   "EMS".Carrier[78].SDC_OUT.HeartBeat := "Clock_1Hz";
   "EMS".Carrier[79].SDC_OUT.HeartBeat := "Clock_1Hz";
   "EMS".Carrier[80].SDC_OUT.HeartBeat := "Clock_1Hz";
END_REGION

REGION Network 2
   // **********************************************************************************************************************
   // 
   // Carrier 71 I-Device Data Transfer Interlocks from Carrier to SDC
   // 
   // **********************************************************************************************************************
   RUNG wire#powerrail
      Coil( "SectionComment" )
   END_RUNG
   // the same network as SCL:
   "SectionComment" := TRUE;
END_REGION

REGION Network 3
   RUNG wire#powerrail
      Contact( "Carrier_71_Status.0" )
      Coil( "EMS".Carrier[71].SDC_IN.HeartBeat )
   END_RUNG
   // the same network as SCL:
   "EMS".Carrier[71].SDC_IN.HeartBeat := "Carrier_71_Status.0";
END_REGION

REGION Network 4
   "C71_Heartbeat_On_Timer".TON(IN := "EMS".Carrier[71].SDC_IN.HeartBeat, PT := T#3s);
END_REGION

REGION Network 5
   "C71_Heartbeat_Off_Timer".TON(IN := NOT "EMS".Carrier[71].SDC_IN.HeartBeat, PT := T#3s);
END_REGION

REGION Network 6
   RUNG wire#powerrail
      Contact( "Carrier_71_Status.7" )
      wire#w1
      Coil( "EMS".Carrier[71].CommFlt )
   END_RUNG
   RUNG wire#powerrail
      Contact( "C71_Heartbeat_On_Timer".Q )
   END_RUNG wire#w1
   RUNG wire#powerrail
      Contact( "C71_Heartbeat_Off_Timer".Q )
   END_RUNG wire#w1
   // the same network as SCL:
   "EMS".Carrier[71].CommFlt := "Carrier_71_Status.7" OR "C71_Heartbeat_On_Timer".Q OR "C71_Heartbeat_Off_Timer".Q;
END_REGION

REGION Network 7
   RUNG wire#powerrail
      Contact( "EMS".Carrier[71].CommFlt )
      JumpCoil( C71_Comm_Fault )
   END_RUNG
   // the same network as SCL:
   IF "EMS".Carrier[71].CommFlt THEN GOTO C71_Comm_Fault; END_IF;
END_REGION

REGION Network 8
   RUNG wire#powerrail
      { S7_Templates := "SrcType := Word" } NE_Contact(in1 := "Carrier_71_CarrierNumber", in2 := 0)
      Move(in := "Carrier_71_CarrierNumber", out1 => "EMS".Carrier[71].SDC_IN.CarrierNumber)
   END_RUNG
   // the same network as SCL:
   IF "Carrier_71_CarrierNumber" <> 0 THEN
       "EMS".Carrier[71].SDC_IN.CarrierNumber := "Carrier_71_CarrierNumber";
   END_IF;
END_REGION

REGION Network 9
   RUNG wire#powerrail
      { S7_Templates := "SrcType := DWord" } NE_Contact(in1 := "Carrier_71_CarrierPosition", in2 := 0)
      Move(in := "Carrier_71_CarrierPosition", out1 => "EMS".Carrier[71].SDC_IN.CarrierPosition)
   END_RUNG
   // the same network as SCL:
   IF "Carrier_71_CarrierPosition" <> 0 THEN
       "EMS".Carrier[71].SDC_IN.CarrierPosition := "Carrier_71_CarrierPosition";
   END_IF;
END_REGION

REGION Network 10
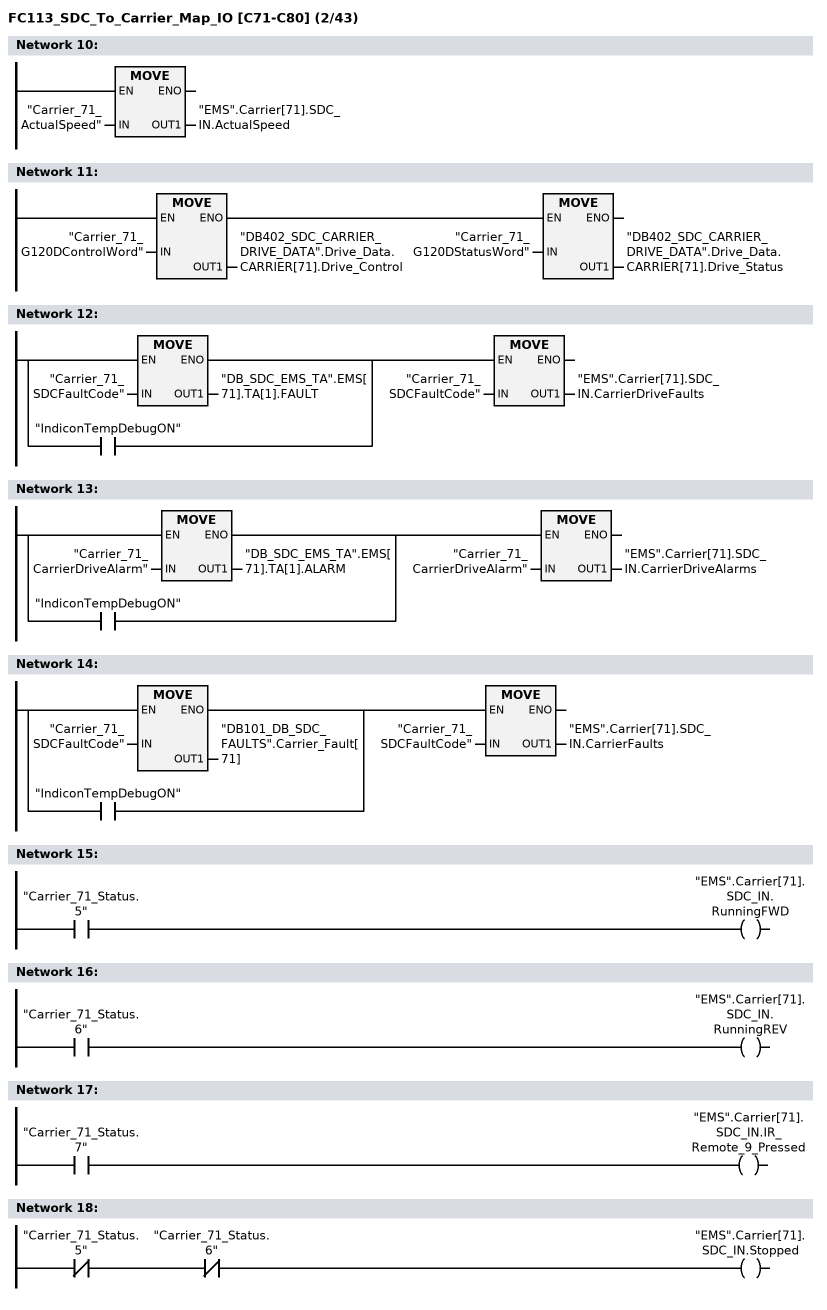
   RUNG wire#powerrail
      Move(in := "Carrier_71_ActualSpeed", out1 => "EMS".Carrier[71].SDC_IN.ActualSpeed)
   END_RUNG
   // the same network as SCL:
   "EMS".Carrier[71].SDC_IN.ActualSpeed := "Carrier_71_ActualSpeed";
END_REGION

REGION Network 11
   RUNG wire#powerrail
      Move(in := "Carrier_71_G120DControlWord", out1 => "DB402_SDC_CARRIER_DRIVE_DATA".Drive_Data.CARRIER[71].Drive_Control)
      Move(in := "Carrier_71_G120DStatusWord", out1 => "DB402_SDC_CARRIER_DRIVE_DATA".Drive_Data.CARRIER[71].Drive_Status)
   END_RUNG
   // the same network as SCL:
   "DB402_SDC_CARRIER_DRIVE_DATA".Drive_Data.CARRIER[71].Drive_Control := "Carrier_71_G120DControlWord";
   "DB402_SDC_CARRIER_DRIVE_DATA".Drive_Data.CARRIER[71].Drive_Status := "Carrier_71_G120DStatusWord";
END_REGION

REGION Network 12
   RUNG wire#powerrail
      Move(in := "Carrier_71_SDCFaultCode", out1 => "DB_SDC_EMS_TA".EMS[71].TA[1].FAULT)
      wire#w1
      Move(in := "Carrier_71_SDCFaultCode", out1 => "EMS".Carrier[71].SDC_IN.CarrierDriveFaults)
   END_RUNG
   RUNG wire#powerrail
      Contact( "IndiconTempDebugON" )
   END_RUNG wire#w1
   // the same network as SCL:
   "DB_SDC_EMS_TA".EMS[71].TA[1].FAULT := "Carrier_71_SDCFaultCode";
   IF TRUE OR "IndiconTempDebugON" THEN
       "EMS".Carrier[71].SDC_IN.CarrierDriveFaults := "Carrier_71_SDCFaultCode";
   END_IF;
END_REGION

REGION Network 13
   RUNG wire#powerrail
      Move(in := "Carrier_71_CarrierDriveAlarm", out1 => "DB_SDC_EMS_TA".EMS[71].TA[1].ALARM)
      wire#w1
      Move(in := "Carrier_71_CarrierDriveAlarm", out1 => "EMS".Carrier[71].SDC_IN.CarrierDriveAlarms)
   END_RUNG
   RUNG wire#powerrail
      Contact( "IndiconTempDebugON" )
   END_RUNG wire#w1
   // the same network as SCL:
   "DB_SDC_EMS_TA".EMS[71].TA[1].ALARM := "Carrier_71_CarrierDriveAlarm";
   IF TRUE OR "IndiconTempDebugON" THEN
       "EMS".Carrier[71].SDC_IN.CarrierDriveAlarms := "Carrier_71_CarrierDriveAlarm";
   END_IF;
END_REGION

REGION Network 14
   RUNG wire#powerrail
      Move(in := "Carrier_71_SDCFaultCode", out1 => "DB101_DB_SDC_FAULTS".Carrier_Fault[71])
      wire#w1
      Move(in := "Carrier_71_SDCFaultCode", out1 => "EMS".Carrier[71].SDC_IN.CarrierFaults)
   END_RUNG
   RUNG wire#powerrail
      Contact( "IndiconTempDebugON" )
   END_RUNG wire#w1
   // the same network as SCL:
   "DB101_DB_SDC_FAULTS".Carrier_Fault[71] := "Carrier_71_SDCFaultCode";
   IF TRUE OR "IndiconTempDebugON" THEN
       "EMS".Carrier[71].SDC_IN.CarrierFaults := "Carrier_71_SDCFaultCode";
   END_IF;
END_REGION

REGION Network 15
   RUNG wire#powerrail
      Contact( "Carrier_71_Status.5" )
      Coil( "EMS".Carrier[71].SDC_IN.RunningFWD )
   END_RUNG
   // the same network as SCL:
   "EMS".Carrier[71].SDC_IN.RunningFWD := "Carrier_71_Status.5";
END_REGION

REGION Network 16
   RUNG wire#powerrail
      Contact( "Carrier_71_Status.6" )
      Coil( "EMS".Carrier[71].SDC_IN.RunningREV )
   END_RUNG
   // the same network as SCL:
   "EMS".Carrier[71].SDC_IN.RunningREV := "Carrier_71_Status.6";
END_REGION

REGION Network 17
   RUNG wire#powerrail
      Contact( "Carrier_71_Status.7" )
      Coil( "EMS".Carrier[71].SDC_IN.IR_Remote_9_Pressed )
   END_RUNG
   // the same network as SCL:
   "EMS".Carrier[71].SDC_IN.IR_Remote_9_Pressed := "Carrier_71_Status.7";
END_REGION

REGION Network 18
   RUNG wire#powerrail
      I_Contact( "Carrier_71_Status.5" )
      I_Contact( "Carrier_71_Status.6" )
      Coil( "EMS".Carrier[71].SDC_IN.Stopped )
   END_RUNG
   // the same network as SCL:
   "EMS".Carrier[71].SDC_IN.Stopped := NOT "Carrier_71_Status.5" AND NOT "Carrier_71_Status.6";
END_REGION

REGION Network 19
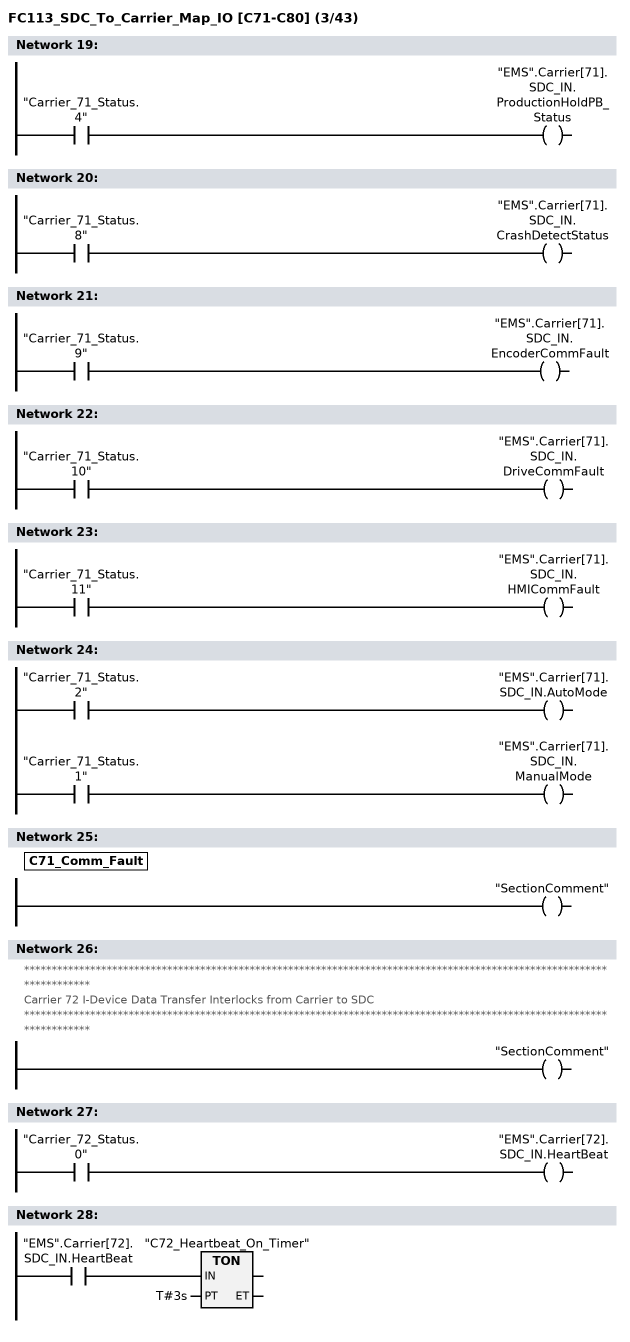
   RUNG wire#powerrail
      Contact( "Carrier_71_Status.4" )
      Coil( "EMS".Carrier[71].SDC_IN.ProductionHoldPB_Status )
   END_RUNG
   // the same network as SCL:
   "EMS".Carrier[71].SDC_IN.ProductionHoldPB_Status := "Carrier_71_Status.4";
END_REGION

REGION Network 20
   RUNG wire#powerrail
      Contact( "Carrier_71_Status.8" )
      Coil( "EMS".Carrier[71].SDC_IN.CrashDetectStatus )
   END_RUNG
   // the same network as SCL:
   "EMS".Carrier[71].SDC_IN.CrashDetectStatus := "Carrier_71_Status.8";
END_REGION

REGION Network 21
   RUNG wire#powerrail
      Contact( "Carrier_71_Status.9" )
      Coil( "EMS".Carrier[71].SDC_IN.EncoderCommFault )
   END_RUNG
   // the same network as SCL:
   "EMS".Carrier[71].SDC_IN.EncoderCommFault := "Carrier_71_Status.9";
END_REGION

REGION Network 22
   RUNG wire#powerrail
      Contact( "Carrier_71_Status.10" )
      Coil( "EMS".Carrier[71].SDC_IN.DriveCommFault )
   END_RUNG
   // the same network as SCL:
   "EMS".Carrier[71].SDC_IN.DriveCommFault := "Carrier_71_Status.10";
END_REGION

REGION Network 23
   RUNG wire#powerrail
      Contact( "Carrier_71_Status.11" )
      Coil( "EMS".Carrier[71].SDC_IN.HMICommFault )
   END_RUNG
   // the same network as SCL:
   "EMS".Carrier[71].SDC_IN.HMICommFault := "Carrier_71_Status.11";
END_REGION

REGION Network 24
   RUNG wire#powerrail
      Contact( "Carrier_71_Status.2" )
      Coil( "EMS".Carrier[71].SDC_IN.AutoMode )
   END_RUNG
   RUNG wire#powerrail
      Contact( "Carrier_71_Status.1" )
      Coil( "EMS".Carrier[71].SDC_IN.ManualMode )
   END_RUNG
   // the same network as SCL:
   "EMS".Carrier[71].SDC_IN.AutoMode := "Carrier_71_Status.2";
   "EMS".Carrier[71].SDC_IN.ManualMode := "Carrier_71_Status.1";
END_REGION

REGION Network 25
   Label( C71_Comm_Fault )
   RUNG wire#powerrail
      Coil( "SectionComment" )
   END_RUNG
   // the same network as SCL:
   C71_Comm_Fault:
   "SectionComment" := TRUE;
END_REGION

REGION Network 26
   // **********************************************************************************************************************
   // 
   // Carrier 72 I-Device Data Transfer Interlocks from Carrier to SDC
   // 
   // **********************************************************************************************************************
   RUNG wire#powerrail
      Coil( "SectionComment" )
   END_RUNG
   // the same network as SCL:
   "SectionComment" := TRUE;
END_REGION

REGION Network 27
   RUNG wire#powerrail
      Contact( "Carrier_72_Status.0" )
      Coil( "EMS".Carrier[72].SDC_IN.HeartBeat )
   END_RUNG
   // the same network as SCL:
   "EMS".Carrier[72].SDC_IN.HeartBeat := "Carrier_72_Status.0";
END_REGION

REGION Network 28
   "C72_Heartbeat_On_Timer".TON(IN := "EMS".Carrier[72].SDC_IN.HeartBeat, PT := T#3s);
END_REGION

REGION Network 29
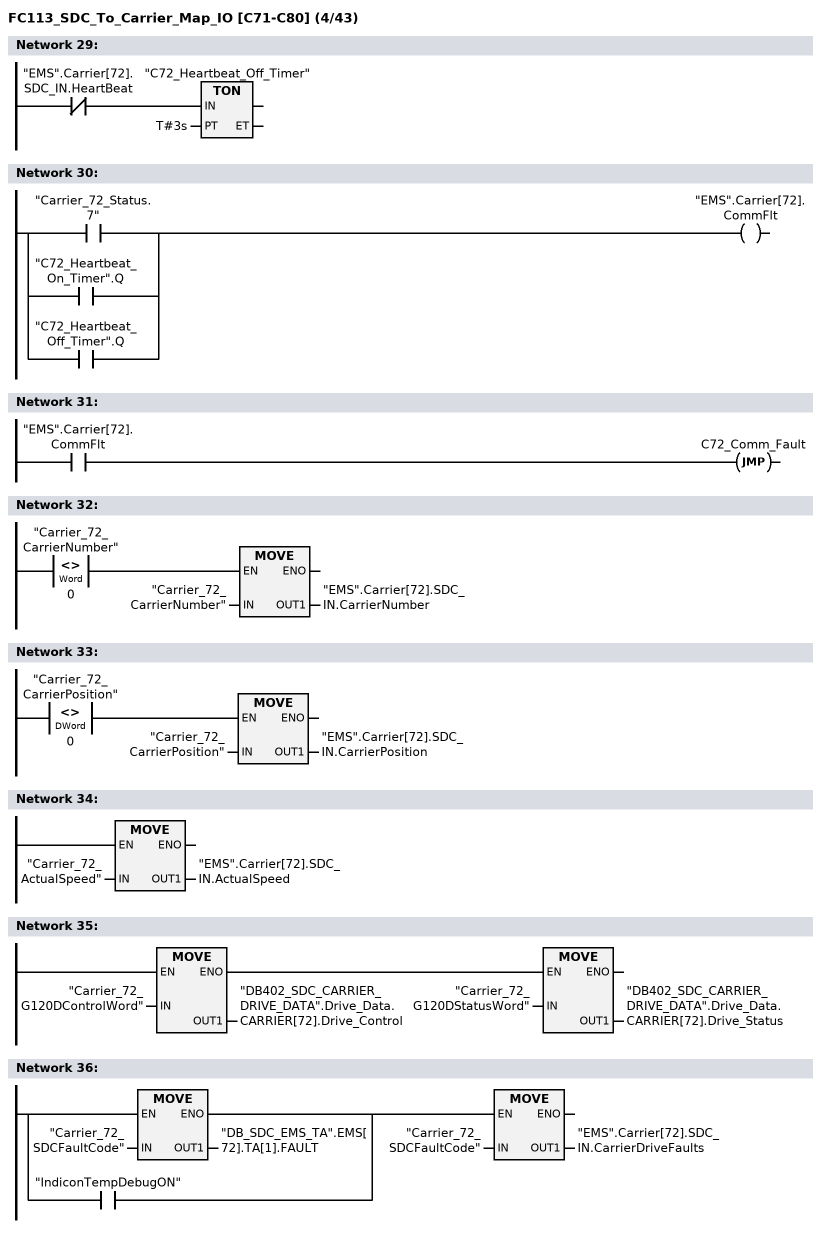
   "C72_Heartbeat_Off_Timer".TON(IN := NOT "EMS".Carrier[72].SDC_IN.HeartBeat, PT := T#3s);
END_REGION

REGION Network 30
   RUNG wire#powerrail
      Contact( "Carrier_72_Status.7" )
      wire#w1
      Coil( "EMS".Carrier[72].CommFlt )
   END_RUNG
   RUNG wire#powerrail
      Contact( "C72_Heartbeat_On_Timer".Q )
   END_RUNG wire#w1
   RUNG wire#powerrail
      Contact( "C72_Heartbeat_Off_Timer".Q )
   END_RUNG wire#w1
   // the same network as SCL:
   "EMS".Carrier[72].CommFlt := "Carrier_72_Status.7" OR "C72_Heartbeat_On_Timer".Q OR "C72_Heartbeat_Off_Timer".Q;
END_REGION

REGION Network 31
   RUNG wire#powerrail
      Contact( "EMS".Carrier[72].CommFlt )
      JumpCoil( C72_Comm_Fault )
   END_RUNG
   // the same network as SCL:
   IF "EMS".Carrier[72].CommFlt THEN GOTO C72_Comm_Fault; END_IF;
END_REGION

REGION Network 32
   RUNG wire#powerrail
      { S7_Templates := "SrcType := Word" } NE_Contact(in1 := "Carrier_72_CarrierNumber", in2 := 0)
      Move(in := "Carrier_72_CarrierNumber", out1 => "EMS".Carrier[72].SDC_IN.CarrierNumber)
   END_RUNG
   // the same network as SCL:
   IF "Carrier_72_CarrierNumber" <> 0 THEN
       "EMS".Carrier[72].SDC_IN.CarrierNumber := "Carrier_72_CarrierNumber";
   END_IF;
END_REGION

REGION Network 33
   RUNG wire#powerrail
      { S7_Templates := "SrcType := DWord" } NE_Contact(in1 := "Carrier_72_CarrierPosition", in2 := 0)
      Move(in := "Carrier_72_CarrierPosition", out1 => "EMS".Carrier[72].SDC_IN.CarrierPosition)
   END_RUNG
   // the same network as SCL:
   IF "Carrier_72_CarrierPosition" <> 0 THEN
       "EMS".Carrier[72].SDC_IN.CarrierPosition := "Carrier_72_CarrierPosition";
   END_IF;
END_REGION

REGION Network 34
   RUNG wire#powerrail
      Move(in := "Carrier_72_ActualSpeed", out1 => "EMS".Carrier[72].SDC_IN.ActualSpeed)
   END_RUNG
   // the same network as SCL:
   "EMS".Carrier[72].SDC_IN.ActualSpeed := "Carrier_72_ActualSpeed";
END_REGION

REGION Network 35
   RUNG wire#powerrail
      Move(in := "Carrier_72_G120DControlWord", out1 => "DB402_SDC_CARRIER_DRIVE_DATA".Drive_Data.CARRIER[72].Drive_Control)
      Move(in := "Carrier_72_G120DStatusWord", out1 => "DB402_SDC_CARRIER_DRIVE_DATA".Drive_Data.CARRIER[72].Drive_Status)
   END_RUNG
   // the same network as SCL:
   "DB402_SDC_CARRIER_DRIVE_DATA".Drive_Data.CARRIER[72].Drive_Control := "Carrier_72_G120DControlWord";
   "DB402_SDC_CARRIER_DRIVE_DATA".Drive_Data.CARRIER[72].Drive_Status := "Carrier_72_G120DStatusWord";
END_REGION

REGION Network 36
   RUNG wire#powerrail
      Move(in := "Carrier_72_SDCFaultCode", out1 => "DB_SDC_EMS_TA".EMS[72].TA[1].FAULT)
      wire#w1
      Move(in := "Carrier_72_SDCFaultCode", out1 => "EMS".Carrier[72].SDC_IN.CarrierDriveFaults)
   END_RUNG
   RUNG wire#powerrail
      Contact( "IndiconTempDebugON" )
   END_RUNG wire#w1
   // the same network as SCL:
   "DB_SDC_EMS_TA".EMS[72].TA[1].FAULT := "Carrier_72_SDCFaultCode";
   IF TRUE OR "IndiconTempDebugON" THEN
       "EMS".Carrier[72].SDC_IN.CarrierDriveFaults := "Carrier_72_SDCFaultCode";
   END_IF;
END_REGION

REGION Network 37
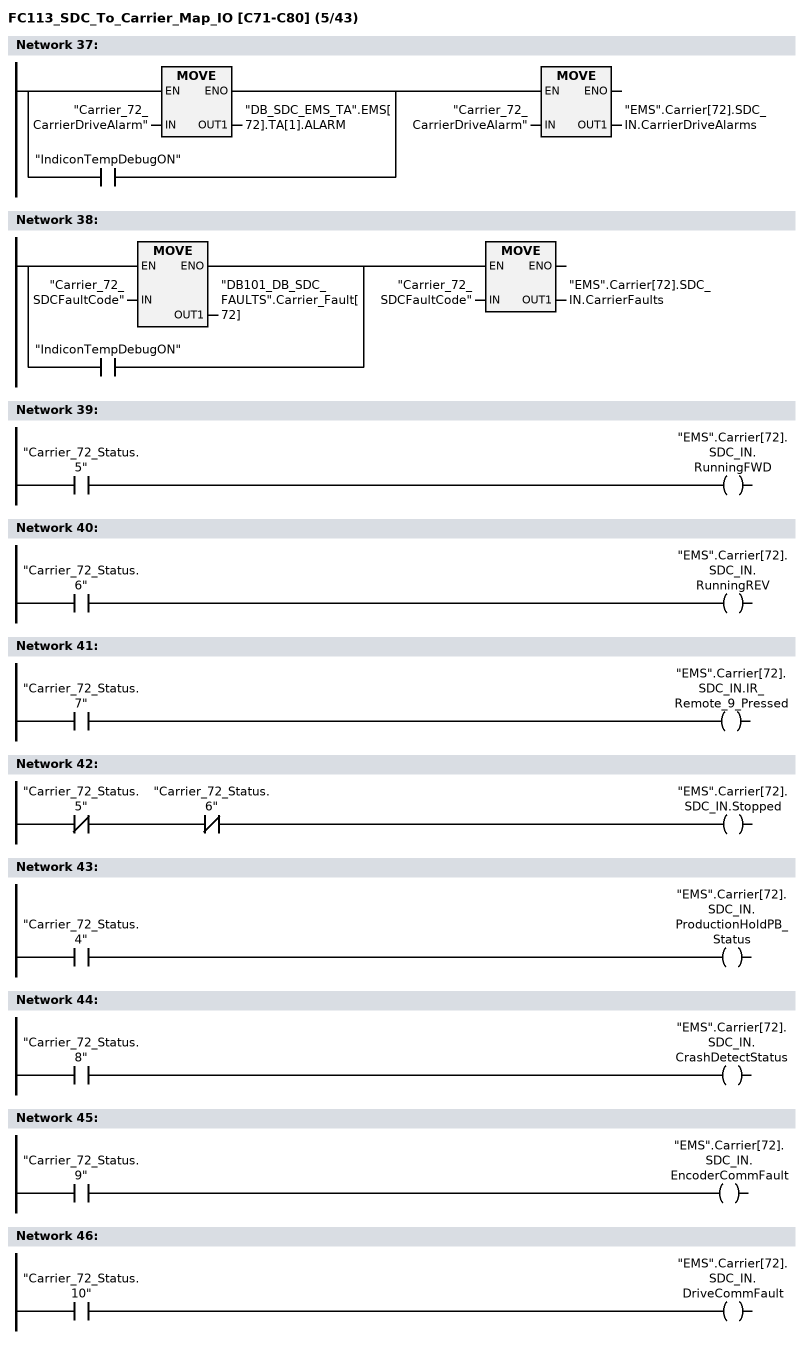
   RUNG wire#powerrail
      Move(in := "Carrier_72_CarrierDriveAlarm", out1 => "DB_SDC_EMS_TA".EMS[72].TA[1].ALARM)
      wire#w1
      Move(in := "Carrier_72_CarrierDriveAlarm", out1 => "EMS".Carrier[72].SDC_IN.CarrierDriveAlarms)
   END_RUNG
   RUNG wire#powerrail
      Contact( "IndiconTempDebugON" )
   END_RUNG wire#w1
   // the same network as SCL:
   "DB_SDC_EMS_TA".EMS[72].TA[1].ALARM := "Carrier_72_CarrierDriveAlarm";
   IF TRUE OR "IndiconTempDebugON" THEN
       "EMS".Carrier[72].SDC_IN.CarrierDriveAlarms := "Carrier_72_CarrierDriveAlarm";
   END_IF;
END_REGION

REGION Network 38
   RUNG wire#powerrail
      Move(in := "Carrier_72_SDCFaultCode", out1 => "DB101_DB_SDC_FAULTS".Carrier_Fault[72])
      wire#w1
      Move(in := "Carrier_72_SDCFaultCode", out1 => "EMS".Carrier[72].SDC_IN.CarrierFaults)
   END_RUNG
   RUNG wire#powerrail
      Contact( "IndiconTempDebugON" )
   END_RUNG wire#w1
   // the same network as SCL:
   "DB101_DB_SDC_FAULTS".Carrier_Fault[72] := "Carrier_72_SDCFaultCode";
   IF TRUE OR "IndiconTempDebugON" THEN
       "EMS".Carrier[72].SDC_IN.CarrierFaults := "Carrier_72_SDCFaultCode";
   END_IF;
END_REGION

REGION Network 39
   RUNG wire#powerrail
      Contact( "Carrier_72_Status.5" )
      Coil( "EMS".Carrier[72].SDC_IN.RunningFWD )
   END_RUNG
   // the same network as SCL:
   "EMS".Carrier[72].SDC_IN.RunningFWD := "Carrier_72_Status.5";
END_REGION

REGION Network 40
   RUNG wire#powerrail
      Contact( "Carrier_72_Status.6" )
      Coil( "EMS".Carrier[72].SDC_IN.RunningREV )
   END_RUNG
   // the same network as SCL:
   "EMS".Carrier[72].SDC_IN.RunningREV := "Carrier_72_Status.6";
END_REGION

REGION Network 41
   RUNG wire#powerrail
      Contact( "Carrier_72_Status.7" )
      Coil( "EMS".Carrier[72].SDC_IN.IR_Remote_9_Pressed )
   END_RUNG
   // the same network as SCL:
   "EMS".Carrier[72].SDC_IN.IR_Remote_9_Pressed := "Carrier_72_Status.7";
END_REGION

REGION Network 42
   RUNG wire#powerrail
      I_Contact( "Carrier_72_Status.5" )
      I_Contact( "Carrier_72_Status.6" )
      Coil( "EMS".Carrier[72].SDC_IN.Stopped )
   END_RUNG
   // the same network as SCL:
   "EMS".Carrier[72].SDC_IN.Stopped := NOT "Carrier_72_Status.5" AND NOT "Carrier_72_Status.6";
END_REGION

REGION Network 43
   RUNG wire#powerrail
      Contact( "Carrier_72_Status.4" )
      Coil( "EMS".Carrier[72].SDC_IN.ProductionHoldPB_Status )
   END_RUNG
   // the same network as SCL:
   "EMS".Carrier[72].SDC_IN.ProductionHoldPB_Status := "Carrier_72_Status.4";
END_REGION

REGION Network 44
   RUNG wire#powerrail
      Contact( "Carrier_72_Status.8" )
      Coil( "EMS".Carrier[72].SDC_IN.CrashDetectStatus )
   END_RUNG
   // the same network as SCL:
   "EMS".Carrier[72].SDC_IN.CrashDetectStatus := "Carrier_72_Status.8";
END_REGION

REGION Network 45
   RUNG wire#powerrail
      Contact( "Carrier_72_Status.9" )
      Coil( "EMS".Carrier[72].SDC_IN.EncoderCommFault )
   END_RUNG
   // the same network as SCL:
   "EMS".Carrier[72].SDC_IN.EncoderCommFault := "Carrier_72_Status.9";
END_REGION

REGION Network 46
   RUNG wire#powerrail
      Contact( "Carrier_72_Status.10" )
      Coil( "EMS".Carrier[72].SDC_IN.DriveCommFault )
   END_RUNG
   // the same network as SCL:
   "EMS".Carrier[72].SDC_IN.DriveCommFault := "Carrier_72_Status.10";
END_REGION

REGION Network 47
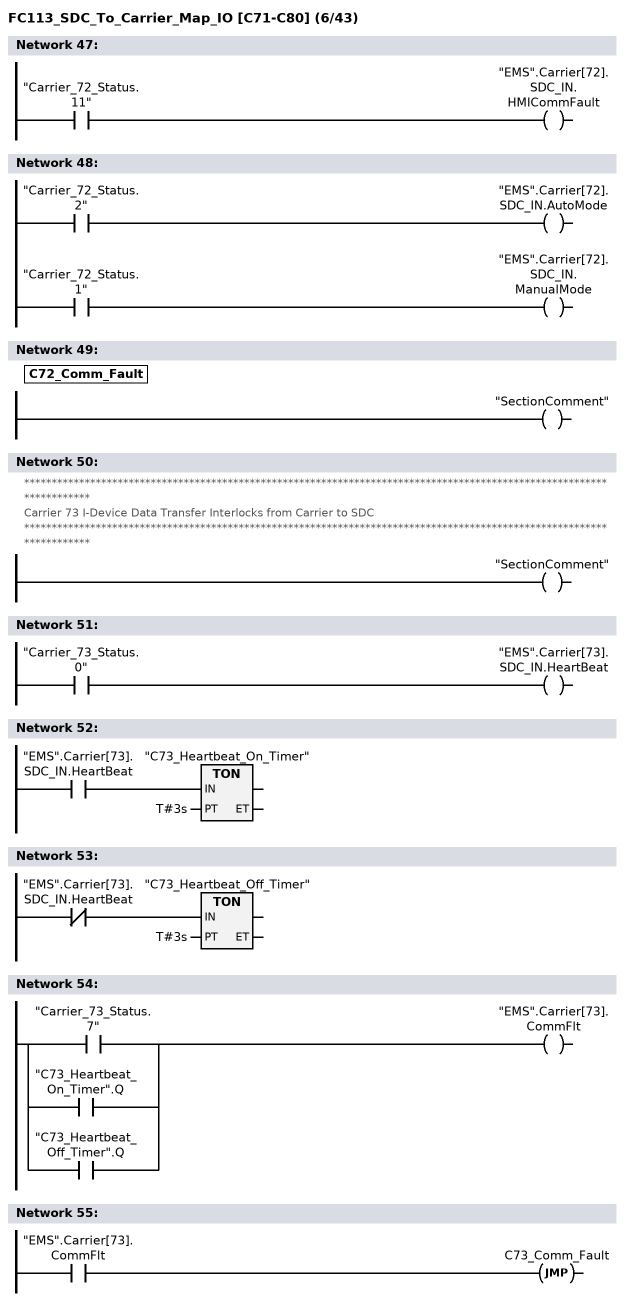
   RUNG wire#powerrail
      Contact( "Carrier_72_Status.11" )
      Coil( "EMS".Carrier[72].SDC_IN.HMICommFault )
   END_RUNG
   // the same network as SCL:
   "EMS".Carrier[72].SDC_IN.HMICommFault := "Carrier_72_Status.11";
END_REGION

REGION Network 48
   RUNG wire#powerrail
      Contact( "Carrier_72_Status.2" )
      Coil( "EMS".Carrier[72].SDC_IN.AutoMode )
   END_RUNG
   RUNG wire#powerrail
      Contact( "Carrier_72_Status.1" )
      Coil( "EMS".Carrier[72].SDC_IN.ManualMode )
   END_RUNG
   // the same network as SCL:
   "EMS".Carrier[72].SDC_IN.AutoMode := "Carrier_72_Status.2";
   "EMS".Carrier[72].SDC_IN.ManualMode := "Carrier_72_Status.1";
END_REGION

REGION Network 49
   Label( C72_Comm_Fault )
   RUNG wire#powerrail
      Coil( "SectionComment" )
   END_RUNG
   // the same network as SCL:
   C72_Comm_Fault:
   "SectionComment" := TRUE;
END_REGION

REGION Network 50
   // **********************************************************************************************************************
   // 
   // Carrier 73 I-Device Data Transfer Interlocks from Carrier to SDC
   // 
   // **********************************************************************************************************************
   RUNG wire#powerrail
      Coil( "SectionComment" )
   END_RUNG
   // the same network as SCL:
   "SectionComment" := TRUE;
END_REGION

REGION Network 51
   RUNG wire#powerrail
      Contact( "Carrier_73_Status.0" )
      Coil( "EMS".Carrier[73].SDC_IN.HeartBeat )
   END_RUNG
   // the same network as SCL:
   "EMS".Carrier[73].SDC_IN.HeartBeat := "Carrier_73_Status.0";
END_REGION

REGION Network 52
   "C73_Heartbeat_On_Timer".TON(IN := "EMS".Carrier[73].SDC_IN.HeartBeat, PT := T#3s);
END_REGION

REGION Network 53
   "C73_Heartbeat_Off_Timer".TON(IN := NOT "EMS".Carrier[73].SDC_IN.HeartBeat, PT := T#3s);
END_REGION

REGION Network 54
   RUNG wire#powerrail
      Contact( "Carrier_73_Status.7" )
      wire#w1
      Coil( "EMS".Carrier[73].CommFlt )
   END_RUNG
   RUNG wire#powerrail
      Contact( "C73_Heartbeat_On_Timer".Q )
   END_RUNG wire#w1
   RUNG wire#powerrail
      Contact( "C73_Heartbeat_Off_Timer".Q )
   END_RUNG wire#w1
   // the same network as SCL:
   "EMS".Carrier[73].CommFlt := "Carrier_73_Status.7" OR "C73_Heartbeat_On_Timer".Q OR "C73_Heartbeat_Off_Timer".Q;
END_REGION

REGION Network 55
   RUNG wire#powerrail
      Contact( "EMS".Carrier[73].CommFlt )
      JumpCoil( C73_Comm_Fault )
   END_RUNG
   // the same network as SCL:
   IF "EMS".Carrier[73].CommFlt THEN GOTO C73_Comm_Fault; END_IF;
END_REGION

REGION Network 56
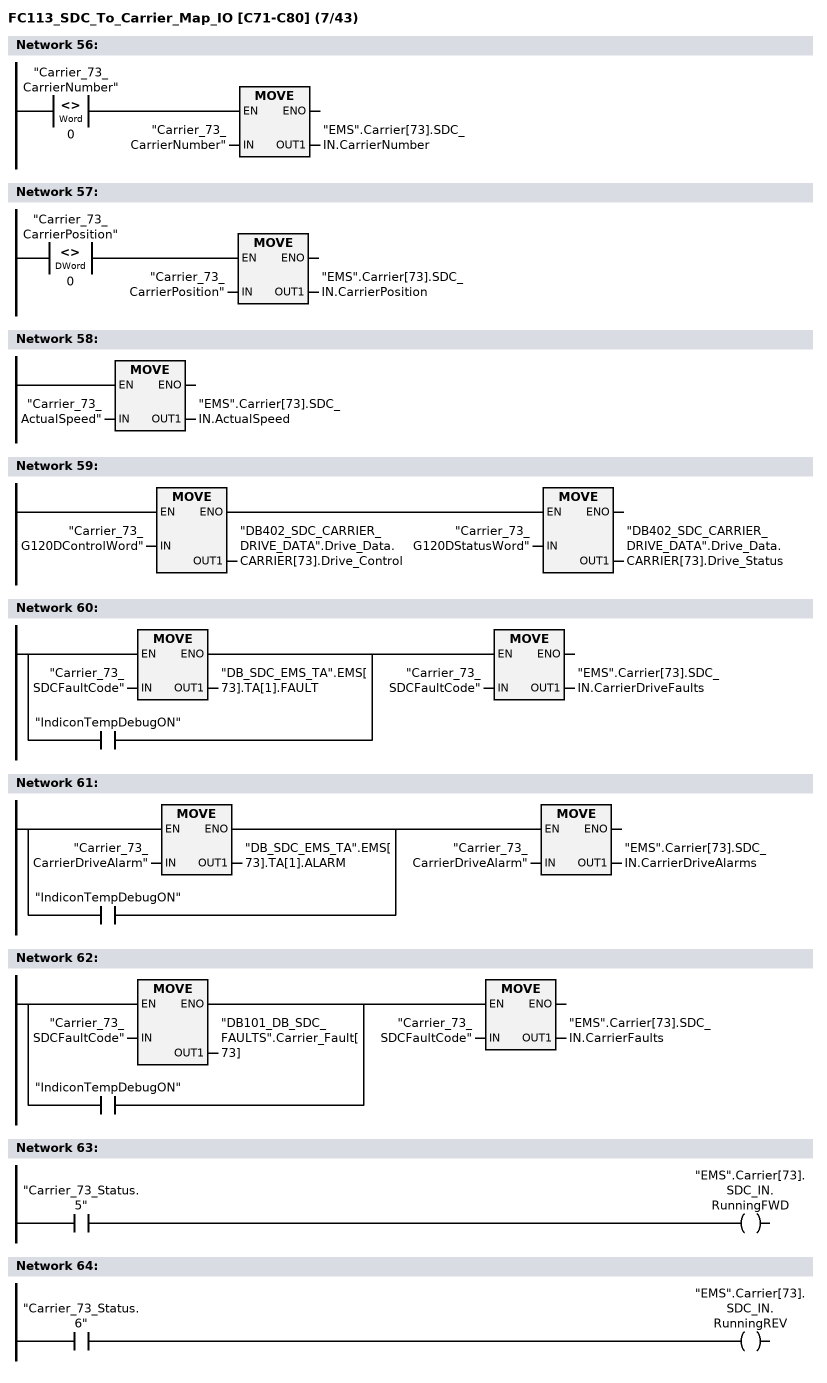
   RUNG wire#powerrail
      { S7_Templates := "SrcType := Word" } NE_Contact(in1 := "Carrier_73_CarrierNumber", in2 := 0)
      Move(in := "Carrier_73_CarrierNumber", out1 => "EMS".Carrier[73].SDC_IN.CarrierNumber)
   END_RUNG
   // the same network as SCL:
   IF "Carrier_73_CarrierNumber" <> 0 THEN
       "EMS".Carrier[73].SDC_IN.CarrierNumber := "Carrier_73_CarrierNumber";
   END_IF;
END_REGION

REGION Network 57
   RUNG wire#powerrail
      { S7_Templates := "SrcType := DWord" } NE_Contact(in1 := "Carrier_73_CarrierPosition", in2 := 0)
      Move(in := "Carrier_73_CarrierPosition", out1 => "EMS".Carrier[73].SDC_IN.CarrierPosition)
   END_RUNG
   // the same network as SCL:
   IF "Carrier_73_CarrierPosition" <> 0 THEN
       "EMS".Carrier[73].SDC_IN.CarrierPosition := "Carrier_73_CarrierPosition";
   END_IF;
END_REGION

REGION Network 58
   RUNG wire#powerrail
      Move(in := "Carrier_73_ActualSpeed", out1 => "EMS".Carrier[73].SDC_IN.ActualSpeed)
   END_RUNG
   // the same network as SCL:
   "EMS".Carrier[73].SDC_IN.ActualSpeed := "Carrier_73_ActualSpeed";
END_REGION

REGION Network 59
   RUNG wire#powerrail
      Move(in := "Carrier_73_G120DControlWord", out1 => "DB402_SDC_CARRIER_DRIVE_DATA".Drive_Data.CARRIER[73].Drive_Control)
      Move(in := "Carrier_73_G120DStatusWord", out1 => "DB402_SDC_CARRIER_DRIVE_DATA".Drive_Data.CARRIER[73].Drive_Status)
   END_RUNG
   // the same network as SCL:
   "DB402_SDC_CARRIER_DRIVE_DATA".Drive_Data.CARRIER[73].Drive_Control := "Carrier_73_G120DControlWord";
   "DB402_SDC_CARRIER_DRIVE_DATA".Drive_Data.CARRIER[73].Drive_Status := "Carrier_73_G120DStatusWord";
END_REGION

REGION Network 60
   RUNG wire#powerrail
      Move(in := "Carrier_73_SDCFaultCode", out1 => "DB_SDC_EMS_TA".EMS[73].TA[1].FAULT)
      wire#w1
      Move(in := "Carrier_73_SDCFaultCode", out1 => "EMS".Carrier[73].SDC_IN.CarrierDriveFaults)
   END_RUNG
   RUNG wire#powerrail
      Contact( "IndiconTempDebugON" )
   END_RUNG wire#w1
   // the same network as SCL:
   "DB_SDC_EMS_TA".EMS[73].TA[1].FAULT := "Carrier_73_SDCFaultCode";
   IF TRUE OR "IndiconTempDebugON" THEN
       "EMS".Carrier[73].SDC_IN.CarrierDriveFaults := "Carrier_73_SDCFaultCode";
   END_IF;
END_REGION

REGION Network 61
   RUNG wire#powerrail
      Move(in := "Carrier_73_CarrierDriveAlarm", out1 => "DB_SDC_EMS_TA".EMS[73].TA[1].ALARM)
      wire#w1
      Move(in := "Carrier_73_CarrierDriveAlarm", out1 => "EMS".Carrier[73].SDC_IN.CarrierDriveAlarms)
   END_RUNG
   RUNG wire#powerrail
      Contact( "IndiconTempDebugON" )
   END_RUNG wire#w1
   // the same network as SCL:
   "DB_SDC_EMS_TA".EMS[73].TA[1].ALARM := "Carrier_73_CarrierDriveAlarm";
   IF TRUE OR "IndiconTempDebugON" THEN
       "EMS".Carrier[73].SDC_IN.CarrierDriveAlarms := "Carrier_73_CarrierDriveAlarm";
   END_IF;
END_REGION

REGION Network 62
   RUNG wire#powerrail
      Move(in := "Carrier_73_SDCFaultCode", out1 => "DB101_DB_SDC_FAULTS".Carrier_Fault[73])
      wire#w1
      Move(in := "Carrier_73_SDCFaultCode", out1 => "EMS".Carrier[73].SDC_IN.CarrierFaults)
   END_RUNG
   RUNG wire#powerrail
      Contact( "IndiconTempDebugON" )
   END_RUNG wire#w1
   // the same network as SCL:
   "DB101_DB_SDC_FAULTS".Carrier_Fault[73] := "Carrier_73_SDCFaultCode";
   IF TRUE OR "IndiconTempDebugON" THEN
       "EMS".Carrier[73].SDC_IN.CarrierFaults := "Carrier_73_SDCFaultCode";
   END_IF;
END_REGION

REGION Network 63
   RUNG wire#powerrail
      Contact( "Carrier_73_Status.5" )
      Coil( "EMS".Carrier[73].SDC_IN.RunningFWD )
   END_RUNG
   // the same network as SCL:
   "EMS".Carrier[73].SDC_IN.RunningFWD := "Carrier_73_Status.5";
END_REGION

REGION Network 64
   RUNG wire#powerrail
      Contact( "Carrier_73_Status.6" )
      Coil( "EMS".Carrier[73].SDC_IN.RunningREV )
   END_RUNG
   // the same network as SCL:
   "EMS".Carrier[73].SDC_IN.RunningREV := "Carrier_73_Status.6";
END_REGION

REGION Network 65
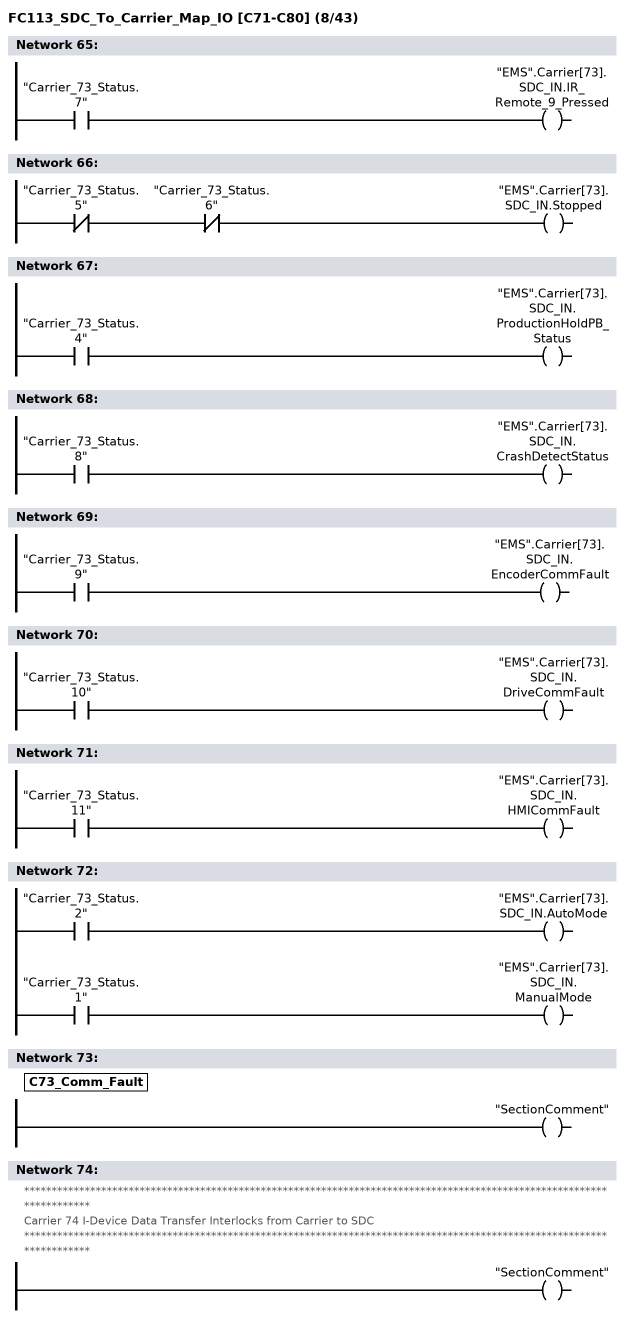
   RUNG wire#powerrail
      Contact( "Carrier_73_Status.7" )
      Coil( "EMS".Carrier[73].SDC_IN.IR_Remote_9_Pressed )
   END_RUNG
   // the same network as SCL:
   "EMS".Carrier[73].SDC_IN.IR_Remote_9_Pressed := "Carrier_73_Status.7";
END_REGION

REGION Network 66
   RUNG wire#powerrail
      I_Contact( "Carrier_73_Status.5" )
      I_Contact( "Carrier_73_Status.6" )
      Coil( "EMS".Carrier[73].SDC_IN.Stopped )
   END_RUNG
   // the same network as SCL:
   "EMS".Carrier[73].SDC_IN.Stopped := NOT "Carrier_73_Status.5" AND NOT "Carrier_73_Status.6";
END_REGION

REGION Network 67
   RUNG wire#powerrail
      Contact( "Carrier_73_Status.4" )
      Coil( "EMS".Carrier[73].SDC_IN.ProductionHoldPB_Status )
   END_RUNG
   // the same network as SCL:
   "EMS".Carrier[73].SDC_IN.ProductionHoldPB_Status := "Carrier_73_Status.4";
END_REGION

REGION Network 68
   RUNG wire#powerrail
      Contact( "Carrier_73_Status.8" )
      Coil( "EMS".Carrier[73].SDC_IN.CrashDetectStatus )
   END_RUNG
   // the same network as SCL:
   "EMS".Carrier[73].SDC_IN.CrashDetectStatus := "Carrier_73_Status.8";
END_REGION

REGION Network 69
   RUNG wire#powerrail
      Contact( "Carrier_73_Status.9" )
      Coil( "EMS".Carrier[73].SDC_IN.EncoderCommFault )
   END_RUNG
   // the same network as SCL:
   "EMS".Carrier[73].SDC_IN.EncoderCommFault := "Carrier_73_Status.9";
END_REGION

REGION Network 70
   RUNG wire#powerrail
      Contact( "Carrier_73_Status.10" )
      Coil( "EMS".Carrier[73].SDC_IN.DriveCommFault )
   END_RUNG
   // the same network as SCL:
   "EMS".Carrier[73].SDC_IN.DriveCommFault := "Carrier_73_Status.10";
END_REGION

REGION Network 71
   RUNG wire#powerrail
      Contact( "Carrier_73_Status.11" )
      Coil( "EMS".Carrier[73].SDC_IN.HMICommFault )
   END_RUNG
   // the same network as SCL:
   "EMS".Carrier[73].SDC_IN.HMICommFault := "Carrier_73_Status.11";
END_REGION

REGION Network 72
   RUNG wire#powerrail
      Contact( "Carrier_73_Status.2" )
      Coil( "EMS".Carrier[73].SDC_IN.AutoMode )
   END_RUNG
   RUNG wire#powerrail
      Contact( "Carrier_73_Status.1" )
      Coil( "EMS".Carrier[73].SDC_IN.ManualMode )
   END_RUNG
   // the same network as SCL:
   "EMS".Carrier[73].SDC_IN.AutoMode := "Carrier_73_Status.2";
   "EMS".Carrier[73].SDC_IN.ManualMode := "Carrier_73_Status.1";
END_REGION

REGION Network 73
   Label( C73_Comm_Fault )
   RUNG wire#powerrail
      Coil( "SectionComment" )
   END_RUNG
   // the same network as SCL:
   C73_Comm_Fault:
   "SectionComment" := TRUE;
END_REGION

REGION Network 74
   // **********************************************************************************************************************
   // 
   // Carrier 74 I-Device Data Transfer Interlocks from Carrier to SDC
   // 
   // **********************************************************************************************************************
   RUNG wire#powerrail
      Coil( "SectionComment" )
   END_RUNG
   // the same network as SCL:
   "SectionComment" := TRUE;
END_REGION

REGION Network 75
